REGION Network 2: Adress_Capa
         L     #Capa_Actual;
         L     1;
         -I;
         L     #Length_Capas;
         *I;
         L     #Offset_Capas;
         +I;
         T     #Adress_Capa;
END_REGION

REGION Network 3: Adress_Filas_DB
   New_Fil:NOP   0;
         L     #Índice_Filas;
         L     1;
         -I;
         L     #Length_Filas_DB;
         *I;
         L     #Offset_Filas_DB;
         +I;
         L     #Adress_Capa;
         +I;
         SLD   3;
         T     #Adress_Filas_DB_bit;
END_REGION

REGION Network 4: Adress_Filas_DI
         L     #Índice_Filas;
         L     1;
         -I;
         L     #Length_Filas_DI;
         *I;
         L     #Offset_Filas_DI;
         +I;
         T     #Adress_Filas_DI;
END_REGION

REGION Network 5: Adress_Elementos_DB
   New_Ele:NOP   0;
         L     #Índice_Elementos;
         L     1;
         -I;
         L     #Length_Elementos_DB_bit;
         *I;
         L     #Offset_Elementos_DB_bit;
         +I;
         L     #Adress_Filas_DB_bit;
         +I;
         T     #Adress_Elementos_DB_bit;
END_REGION

REGION Network 6: Adress_Elementos_DI
         L     #Índice_Elementos;
         L     1;
         -I;
         L     #Length_Elementos_DI;
         *I;
         L     #Offset_Elementos_DI;
         +I;
         L     #Adress_Filas_DI;
         +I;
         T     #Adress_Elementos_DI;
END_REGION

REGION Network 7: AR1 y AR2
         L     #Adress_Elementos_DB_bit;
         LAR1;
         L     #Adress_Elementos_DI;
         SLD   3;
         LAR2;
END_REGION

REGION Network 8: Transferencia de Figuras
   // No debería entrar nunca en este segmento, ya que necesita a Editando_Recetas y no entraría al bloque
         A     "Editando_Recetas";
         AN    "flanco"."nHMI.Pls_Inc_Capa";
         AN    "flanco"."nHMI.Pls_Dec_Capa";
         JCN   Fin;
         OPN   "DB_Receta_Actual";
         OPNDI "DB_Animación";
   // 0 = Invisible
   // 1 = V
   // 2 = H
   // 3 = HH
   //... Creo...
         L     DIB [ AR2 , P#0.0 ];
         L     0;
         ==I;
         JCN   NO_00;
         R     DBX[AR1,P#0.0];
         R     DBX [ AR1 , P#2.0 ];
         JU    Fin;
   NO_00:L     DIB [ AR2 , P#0.0 ];
         L     1;
         ==I;
         JCN   NO_10;
         S     DBX [ AR1 , P#0.0 ];
         R     DBX [ AR1 , P#2.0 ];
         JU    Fin;
   NO_10:L     DIB [ AR2 , P#0.0 ];
         L     2;
         ==I;
         JCN   NO_20;
         R     DBX[AR1,P#0.0];
         S     DBX [ AR1 , P#2.0 ];
         JU    Fin;
   NO_20:S     DBX [ AR1 , P#0.0 ];
         S     DBX [ AR1 , P#2.0 ];
   Fin:  NOP   0;
END_REGION

REGION Network 9: Transferencia de Figuras
   // En base a las figuras en bits de la receta actual, dibuja la capa gráficamente.
         OPN   "DB_Receta_Actual";
         OPNDI "DB_Animación";
   // 0 = Invisible
   // 1 = V
   // 2 = H
   // 3 = HH
   //... Creo...

         AN    DBX [ AR1 , P#0.0 ];
         AN    DBX [ AR1 , P#2.0 ];
         JCN   NO_0;
         L     0;
         JU    Transferir;
   NO_0: A     DBX [ AR1 , P#0.0 ];
         AN    DBX [ AR1 , P#2.0 ];
         JCN   NO_1;
         L     1;
         JU    Transferir;
   NO_1: AN    DBX [ AR1 , P#0.0 ];
         A     DBX [ AR1 , P#2.0 ];
         JCN   NO_2;
         L     2;
         JU    Transferir;
   NO_2: L     3;
   Transferir:T     DIB [ AR2 , P#0.0 ];
END_REGION

REGION Network 10: Transferencia de Elemento_SEL [ Anulado ]
   // Entra a veces en este segmento, se puede pulsar este botón dela pantalla 20 ó 21 [21 no entra al FC]
         A     "flanco"."pHMI.Pls_CargarReceta";
         JCN   Anular;
         OPN   "DB_Receta_Actual";
         OPNDI "DB_Animación";

         SET;
         A     DBX [ AR1 , P#4.0 ];
         JCN   otro;
         L     #Índice_Filas;
         T     "DB_Animación".Fila_SEL;
         L     #Índice_Elementos;
         T     "DB_Animación".Elemento_SEL;
   otro: NOP   0;

   Anular:NOP   0;
         OPN   "DB_Receta_Actual";
         OPNDI "DB_Animación";
END_REGION

REGION Network 11: Bucle Elementos
         L     #Índice_Elementos;
         L     1;
         +I;
         T     #Índice_Elementos;
         L     #Max_Nro_Elementos;
         <=I;
         JC    New_Ele;
END_REGION

REGION Network 12: Bucle Filas
         L     1;
         T     #Índice_Elementos;
         L     #Índice_Filas;
         L     1;
         +I;
         T     #Índice_Filas;
         L     #Max_Nro_Filas;
         <=I;
         JC    New_Fil;
END_REGION

REGION Network 13: Fin de Bloque
         BEU;
END_REGION
END_FUNCTION

FUNCTION "FC_INC_ELEM_ACTUAL" : Void   // FC19, STL
{ S7_Optimized_Access := 'FALSE' }
VERSION : 0.1
BEGIN

REGION Network 1: Constantes
         L     "Proceso Dosificador".Cant_Pallets;
         T     #Nro_Pallet;
         L     "Proceso Dosificador".Capa_Actual;
         T     #Capa_Actual;
         L     38;
         T     #Length_Capas;
         L     54;
         T     #Offset_Capas;
         L     6;
         T     #Length_Filas_DB;
         L     0;
         T     #Offset_Filas_DB;
         L     1;
         T     #Length_Elementos_DB_bit;
         L     0;
         T     #Offset_Elementos_DB_bit;

         L     1;
         T     #Índice_Filas;
         T     #Índice_Elementos;

         L     "Puntero".Max_Nro_Elementos;
         T     #Max_Nro_Elementos;
         L     "Puntero".Max_Nro_Filas;
         T     #Max_Nro_Filas;
         L     "Puntero".Max_Nro_Capas;
         T     #Max_Nro_Capas;
END_REGION

REGION Network 2: Adress_Capa
         L     #Capa_Actual;
         L     1;
         -I;
         L     #Length_Capas;
         *I;
         L     #Offset_Capas;
         +I;
         T     #Adress_Capa;
END_REGION

REGION Network 3: Adress_Filas
   New_Fil:NOP   0;
         L     #Índice_Filas;
         L     1;
         -I;
         L     #Length_Filas_DB;
         *I;
         L     #Offset_Filas_DB;
         +I;
         L     #Adress_Capa;
         +I;
         SLD   3;
         T     #Adress_Filas_DB_bit;
END_REGION

REGION Network 4: Adress_Elementos_DB
   New_Ele:NOP   0;
         L     #Índice_Elementos;
         L     1;
         -I;
         L     #Length_Elementos_DB_bit;
         *I;
         L     #Offset_Elementos_DB_bit;
         +I;
         L     #Adress_Filas_DB_bit;
         +I;
         T     #Adress_Elementos_DB_bit;
END_REGION

REGION Network 5: AR1
         L     #Adress_Elementos_DB_bit;
         LAR1;
END_REGION

REGION Network 6: Habilita ir 1 lugar a la IZQ si gráficamente existe un elemento a la izq.
         OPN   "DB_Receta_Actual";
         SET;
         R     #Habil_1_IZQ;
         L     #Índice_Elementos;
         L     #Max_Nro_Elementos;
         >=I;
         JC    No1IZQ;
         TAR1  AR2;
         L     1;
         +AR2;
         O     DBX [ AR2 , P#0.0 ];
         O     DBX [ AR2 , P#2.0 ];
         =     #Habil_1_IZQ;
   No1IZQ:NOP   0;
END_REGION

REGION Network 7: Habilita ir 2 lugar a la IZQ si gráficamente existen dos elementos a la izq.
         OPN   "DB_Receta_Actual";
         SET;
         R     #Habil_2_IZQ;
         L     #Índice_Elementos;
         L     1;
         +I;
         L     #Max_Nro_Elementos;
         >=I;
         JC    No2IZQ;
         TAR1  AR2;
         L     2;
         +AR2;
         O     DBX [ AR2 , P#0.0 ];
         O     DBX [ AR2 , P#2.0 ];
         =     #Habil_2_IZQ;
   No2IZQ:NOP   0;
END_REGION

REGION Network 8: Habilita ir a ABA_Elem_1 si gráficamente existe el primer elemento de la fila de abajo.
         OPN   "DB_Receta_Actual";
         SET;
         R     #Habil_1_ABA;
         L     #Índice_Filas;
         L     #Max_Nro_Filas;
         >=I;
         JC    No1ABA;
         L     #Adress_Filas_DB_bit;
         SRD   3;
         L     #Length_Filas_DB;
         +I;
         SLD   3;
         L     #Offset_Elementos_DB_bit;
         +I;
         LAR2;
         O     DBX [AR2, P#0.0];
         O     DBX [ AR2 , P#2.0 ];
         =     #Habil_1_ABA;
   No1ABA:NOP   0;
END_REGION

REGION Network 9: Habilita ir a ABA_Elem_2 si gráficamente existe el segundo elemento de la fila de abajo.
         OPN   "DB_Receta_Actual";
         SET;
         R     #Habil_2_ABA;
         L     #Índice_Filas;
         L     #Max_Nro_Filas;
         >=I;
         JC    No2ABA;
         L     #Adress_Filas_DB_bit;
         SRD   3;
         L     #Length_Filas_DB;
         +I;
         SLD   3;
         L     #Offset_Elementos_DB_bit;
         +I;
         L     #Length_Elementos_DB_bit;
         +I;
         LAR2;
         O     DBX [AR2, P#0.0];
         O     DBX [ AR2 , P#2.0 ];
         =     #Habil_2_ABA;
   No2ABA:NOP   0;
END_REGION

REGION Network 10: Habilita cambiar de CAPA_Elem_1, si existe el primer elemento de la próx. capa.
         OPN   "DB_Receta_Actual";
         SET;
         R     #Habil_1_CAPA;
         L     #Capa_Actual;
         L     #Max_Nro_Capas;
         >=I;
         JC    No1CAPA;
         L     #Adress_Capa;
         L     #Length_Capas;
         +I;
         L     #Offset_Filas_DB;
         +I;
         SLD   3;
         L     #Offset_Elementos_DB_bit;
         +I;
         LAR2;
         O     DBX [AR2, P#0.0];
         O     DBX [ AR2 , P#2.0 ];
         =     #Habil_1_CAPA;
   No1CAPA:NOP   0;
END_REGION

REGION Network 11: Habilita cambiar de CAPA_Elem_2, si existe el segundo elemento de la próx. capa.
         OPN   "DB_Receta_Actual";
         SET;
         R     #Habil_2_CAPA;
         L     #Capa_Actual;
         L     #Max_Nro_Capas;
         >=I;
         JC    No2CAPA;
         L     #Adress_Capa;
         L     #Length_Capas;
         +I;
         L     #Offset_Filas_DB;
         +I;
         SLD   3;
         L     #Offset_Elementos_DB_bit;
         +I;
         L     #Length_Elementos_DB_bit;
         +I;
         LAR2;
         O     DBX [AR2, P#0.0];
         O     DBX [ AR2 , P#2.0 ];
         =     #Habil_2_CAPA;
   No2CAPA:NOP   0;
END_REGION

REGION Network 12: #Elemento_Actual
         OPN   "DB_Receta_Actual";

         A     DBX [ AR1 , P#4.0 ];
         =     #Elemento_Actual;

         A     #Elemento_Actual;
         JCN   NoActual;
         TAR1  AR2;
END_REGION

REGION Network 13: NUM = 1
         L     #NUM;
         L     1;
         ==I;
         JCN   NUM_2;
         R     DBX [ AR1 , P#4.0 ];
         A     #Habil_1_IZQ;
         JCN   No_1_IZQ;

         TAR1  AR2;
         L     1;
         +AR2;
         S     DBX [ AR2 , P#4.0 ];
         JU    Fin;

   No_1_IZQ:A     #Habil_1_ABA;
         JCN   No_ABA;
         L     #Adress_Filas_DB_bit;
         SRD   3;
         L     #Length_Filas_DB;
         +I;
         SLD   3;
         L     #Offset_Elementos_DB_bit;
         +I;
         LAR2;
         SET;
         S     DBX [ AR2 , P#4.0 ];
         JU    Fin;

   No_ABA:A     #Habil_1_CAPA;
         JCN   No_CAPA;
         L     #Adress_Capa;
         L     #Length_Capas;
         +I;
         L     #Offset_Filas_DB;
         +I;
         SLD   3;
         L     #Offset_Elementos_DB_bit;
         +I;
         LAR2;
         S     DBX [ AR2 , P#4.0 ];
         L     #Capa_Actual;
         L     1;
         +I;
         T     #Capa_Actual;
         JU    Fin;

   No_CAPA:NOP   0;
         L     #Offset_Capas;
         L     #Offset_Filas_DB;
         +I;
         SLD   3;
         L     #Offset_Elementos_DB_bit;
         +I;
         LAR2;
         S     DBX [ AR2 , P#4.0 ];
         L     1;
         T     #Capa_Actual;
         L     #Nro_Pallet;
         L     1;
         +I;
         T     #Nro_Pallet;
         JU    Fin;
END_REGION

REGION Network 14: NUM = 2
   NUM_2:L     #NUM;
         L     2;
         ==I;
         JCN   NoNUM;
         R     DBX [ AR1 , P#4.0 ];
         A     #Habil_2_IZQ;
         JC    x_2IZQ;
         A     #Habil_1_IZQ;
         A     #Habil_1_ABA;
         JC    x_1IZQ_1ABA;
         A     #Habil_1_IZQ;
         A     #Habil_1_CAPA;
         JC    x_1IZQ_1CAPA;
         A     #Habil_1_IZQ;
         JC    x_1IZQ_1PALLET;
         A     #Habil_2_ABA;
         JC    x_2ABA;
         A     #Habil_1_ABA;
         A     #Habil_1_CAPA;
         JC    x_1ABA_1CAPA;
         A     #Habil_1_ABA;
         JC    x_1ABA_1PALLET;
         A     #Habil_2_CAPA;
         JC    x_2CAPA;
         A     #Habil_1_CAPA;
         JC    x_1CAPA_1PALLET;
         JU    x_2PALLET;

   x_2IZQ:NOP   0;
         TAR1  AR2;
         L     2;
         +AR2;
         S     DBX [ AR2 , P#4.0 ];
         JU    Fin;

   x_1IZQ_1ABA:NOP   0;
         L     #Adress_Filas_DB_bit;
         SRD   3;
         L     #Length_Filas_DB;
         +I;
         SLD   3;
         L     #Offset_Elementos_DB_bit;
         +I;
         LAR2;
         S     DBX [ AR2 , P#4.0 ];
         JU    Fin;

   x_2ABA:NOP   0;
         L     #Adress_Filas_DB_bit;
         SRD   3;
         L     #Length_Filas_DB;
         +I;
         SLD   3;
         L     #Offset_Elementos_DB_bit;
         +I;
         L     #Length_Elementos_DB_bit;
         +I;
         LAR2;
         S     DBX [ AR2 , P#4.0 ];
         JU    Fin;

   x_1IZQ_1CAPA:NOP   0;
   x_1ABA_1CAPA:NOP   0;
         L     #Adress_Capa;
         L     #Length_Capas;
         +I;
         L     #Offset_Filas_DB;
         +I;
         SLD   3;
         L     #Offset_Elementos_DB_bit;
         +I;
         LAR2;
         S     DBX [ AR2 , P#4.0 ];
         L     #Capa_Actual;
         L     1;
         +I;
         T     #Capa_Actual;
         JU    Fin;

   x_2CAPA:NOP   0;
         L     #Adress_Capa;
         L     #Length_Capas;
         +I;
         L     #Offset_Filas_DB;
         +I;
         SLD   3;
         L     #Offset_Elementos_DB_bit;
         +I;
         L     #Length_Elementos_DB_bit;
         +I;
         LAR2;
         S     DBX [ AR2 , P#4.0 ];
         L     #Capa_Actual;
         L     1;
         +I;
         T     #Capa_Actual;
         JU    Fin;

   x_1IZQ_1PALLET:NOP   0;
   x_1ABA_1PALLET:NOP   0;
   x_1CAPA_1PALLET:NOP   0;
         L     #Offset_Capas;
         L     #Offset_Filas_DB;
         +I;
         SLD   3;
         L     #Offset_Elementos_DB_bit;
         +I;
         LAR2;
         S     DBX [ AR2 , P#4.0 ];
         L     1;
         T     #Capa_Actual;
         L     #Nro_Pallet;
         L     1;
         +I;
         T     #Nro_Pallet;
         JU    Fin;

   x_2PALLET:NOP   0;
         L     #Offset_Capas;
         L     #Offset_Filas_DB;
         +I;
         SLD   3;
         L     #Offset_Elementos_DB_bit;
         +I;
         L     #Length_Elementos_DB_bit;
         +I;
         LAR2;
         S     DBX [ AR2 , P#4.0 ];
         L     1;
         T     #Capa_Actual;
         L     #Nro_Pallet;
         L     1;
         +I;
         T     #Nro_Pallet;
         JU    Fin;
END_REGION

REGION Network 15: No elemento actual
   NoNUM:JU    Fin;
   NoActual:NOP   0;
END_REGION

REGION Network 16: Bucle Elementos
         L     #Índice_Elementos;
         L     1;
         +I;
         T     #Índice_Elementos;
         L     #Max_Nro_Elementos;
         <=I;
         JC    New_Ele;
END_REGION

REGION Network 17: Bucle Filas
         L     1;
         T     #Índice_Elementos;
         L     #Índice_Filas;
         L     1;
         +I;
         T     #Índice_Filas;
         L     #Max_Nro_Filas;
         <=I;
         JC    New_Fil;
END_REGION

REGION Network 18: #Error
         SET;
         S     #Error;
         JU    ERROR;
END_REGION

REGION Network 19: Fin de Bloque
   Fin:  SET;
         R     #Error;
         OPN   "DB_Receta_Actual";
         AN    DBX [ AR2 , P#0.0 ];
         AN    DBX [ AR2 , P#2.0 ];
         JCN   NO_0;
         L     0;
         JU    Transferir;
   NO_0: A     DBX [ AR2 , P#0.0 ];
         AN    DBX [ AR2 , P#2.0 ];
         JCN   NO_1;
         L     1;
         JU    Transferir;
   NO_1: AN    DBX [ AR2 , P#0.0 ];
         A     DBX [ AR2 , P#2.0 ];
         JCN   NO_2;
         L     2;
         JU    Transferir;
   NO_2: L     3;
   Transferir:T     "Proceso Dosificador".Elemento_Actual;
   // 0 = Invisible
   // 1 = V
   // 2 = H
   // 3 = HH


   ERROR:L     #Capa_Actual;
         T     "Proceso Dosificador".Capa_Actual;
         L     #Nro_Pallet;
         T     "Proceso Dosificador".Cant_Pallets;
END_REGION
END_FUNCTION

FUNCTION "FC_Ver_Recetas_faltaEditar" : Void   // FC21, STL
TITLE = Muestra los datos de la receta seleccionada
{ S7_Optimized_Access := 'FALSE' }
VERSION : 0.1
BEGIN

REGION Network 1: Constantes
         L     "Puntero".Offset_Recetas;
         T     #Offset_Recetas;
         L     "Puntero".Length_Recetas;
         T     #Length_Recetas;
         L     "Puntero".Offset_Nombre_Receta;
         T     #Offset_Nombre_Receta_DB;
         L     "Puntero".Max_Nro_Recetas;
         T     #Max_Nro_Recetas;
   //
         L     "Puntero".Offset_CapasDist_Receta;
   //    L     51
         T     #Offset_CapasDist_Receta_DB;
         L     "Puntero".Offset_CantCapas_Receta;
   //    L     50
         T     #Offset_CantCapas_Receta_DB;
         L     "Puntero".Length_Nombre_Receta;
   //    L     50
         T     #Length_Nombre_Receta;
   //
         L     316;
         T     #Offset_CantCapas_Receta_DI;
         L     317;
         T     #Offset_CapasDist_Receta_DI;
   //
         L     "DB_Animación".Nro_Receta_Edición;
         T     #Nro_Receta;
   //
         A     "flanco"."nHMI.Pls_Inc_Receta";
         =     #fn_Inc_Receta;
         A     "flanco"."nHMI.Pls_Dec_Receta";
         =     #fn_Dec_Receta;
   //
         L     "HMI".Imagen_Actual;
         T     #Imagen;
END_REGION

REGION Network 2
         L     #Nro_Receta;
         L     #Max_Nro_Recetas;
         <I;
         A     #fn_Inc_Receta;
         JCN   noINC;
         TAK;
         L     1;
         +I;
         JU    Transferir;
   noINC:NOP   0;

         L     #Nro_Receta;
         L     1;
         >I;
         A     #fn_Dec_Receta;
         JCN   noDEC;
         TAK;
         L     1;
         -I;
         JU    Transferir;
   noDEC:NOP   0;
         L     #Nro_Receta;
   Transferir:T     #Nro_Receta;
END_REGION

REGION Network 3: Abrir la receta correspondiente
         L     #Nro_Receta;
         L     1;
         -I;
         L     #Length_Recetas;
         *I;
         L     #Offset_Recetas;
         +I;
         T     #Adress_Receta;
END_REGION

REGION Network 4: Transferir Nombre de receta
         OPN   "DB_RECETAS";
         OPNDI "DB_Animación";
         L     #Adress_Receta;
         L     #Offset_Nombre_Receta_DB;
         +I;
         SLD   3;
         LAR1;
         L     266;
         SLD   3;
         LAR2;
         L     0;
         T     #K;
   Bucle:SLD   3;
         +AR1;
         +AR2;

         A     "Editando_Recetas";
         JCN   NoEsc_0;
         L     DIB [ AR2 , P#0.0 ];
         T     DBB [ AR1 , P#0.0 ];
   NoEsc_0:NOP   0;

         L     DBB [ AR1 , P#0.0 ];
         T     DIB [ AR2 , P#0.0 ];
         L     #K;
         L     1;
         +I;
         T     #K;
         L     #Length_Nombre_Receta;
         <I;
         L     1;
         JC    Bucle;
END_REGION

REGION Network 5: Transferir Número de capas por pallet
         OPN   "DB_RECETAS";
         OPNDI "DB_Animación";
         L     #Adress_Receta;
         L     #Offset_CantCapas_Receta_DB;
         +I;
         SLD   3;
         LAR1;
         L     #Offset_CantCapas_Receta_DI;
         SLD   3;
         LAR2;

         A     "Editando_Recetas";
         JCN   NoEsc_1;
         L     DIB [ AR2 , P#0.0 ];
         T     DBB [ AR1 , P#0.0 ];
   NoEsc_1:NOP   0;

         L     DBB [AR1, P#0.0];
         T     DIB [ AR2 , P#0.0 ];
END_REGION

REGION Network 6: Transferir Número de capas distintas
         OPN   "DB_RECETAS";
         OPNDI "DB_Animación";
         L     #Adress_Receta;
         L     #Offset_CapasDist_Receta_DB;
         +I;
         SLD   3;
         LAR1;
         L     #Offset_CapasDist_Receta_DI;
         SLD   3;
         LAR2;

         A     "Editando_Recetas";
         JCN   NoEsc_2;
         L     DIB [ AR2 , P#0.0 ];
         T     DBB [ AR1 , P#0.0 ];
   NoEsc_2:NOP   0;

         L     DBB [AR1, P#0.0];
         T     DIB [ AR2 , P#0.0 ];
END_REGION

REGION Network 7
         L     #Nro_Receta;
         T     "DB_Animación".Nro_Receta_Edición;
END_REGION
END_FUNCTION

FUNCTION "FC_RESET_ELEM_ACTUAL" : Void   // FC22, STL
{ S7_Optimized_Access := 'FALSE' }
VERSION : 0.1
// Con los datos del dosificador, setea el bit de elemento actual en DB_Receta_Actual
BEGIN

REGION Network 1: Constantes
         L     "Proceso Empujador".Capa_Actual;
         T     #Capa_Empuj;
         L     "Proceso Dosificador".Cant_Pallets;
         T     #Nro_Pallet;
         L     "Proceso Dosificador".Capa_Actual;
         T     #Capa_Actual;
         L     38;
         T     #Length_Capas;
         L     54;
         T     #Offset_Capas;
         L     6;
         T     #Length_Filas_DB;
         L     0;
         T     #Offset_Filas_DB;
         L     1;
         T     #Length_Elementos_DB_bit;
         L     0;
         T     #Offset_Elementos_DB_bit;

         L     1;
         T     #Índice_Capas;
         T     #Índice_Filas;
         T     #Índice_Elementos;

         L     "Puntero".Max_Nro_Elementos;
         T     #Max_Nro_Elementos;
         L     "Puntero".Max_Nro_Filas;
         T     #Max_Nro_Filas;
         L     "Puntero".Max_Nro_Capas;
         T     #Max_Nro_Capas;

         L     "DB_Animación".Fila_SEL;
         T     #Fila_SEL;
         L     "DB_Animación".Elemento_SEL;
         T     #Elemento_SEL;
END_REGION

REGION Network 2: Set CAPA
         OPN   "DB_Receta_Actual";
   //     SPA   no
         L     #Capa_Empuj;
         T     #Capa_Actual;
   no:   NOP   0;
END_REGION

REGION Network 3: Adress_Capa
   New_Cap:L     #Índice_Capas;
         L     1;
         -I;
         L     #Length_Capas;
         *I;
         L     #Offset_Capas;
         +I;
         T     #Adress_Capa;
END_REGION

REGION Network 4: Adress_Filas
   New_Fil:L     #Índice_Filas;
         L     1;
         -I;
         L     #Length_Filas_DB;
         *I;
         L     #Offset_Filas_DB;
         +I;
         L     #Adress_Capa;
         +I;
         SLD   3;
         T     #Adress_Filas_DB_bit;
END_REGION

REGION Network 5: Adress_Elementos_DB
   New_Ele:L     #Índice_Elementos;
         L     1;
         -I;
         L     #Length_Elementos_DB_bit;
         *I;
         L     #Offset_Elementos_DB_bit;
         +I;
         L     #Adress_Filas_DB_bit;
         +I;
         T     #Adress_Elementos_DB_bit;
END_REGION

REGION Network 6: AR1
         L     #Adress_Elementos_DB_bit;
         LAR1;
END_REGION

REGION Network 7: SR Elemento actual
   //  SPA   end
         L     #Capa_Actual;
         L     #Índice_Capas;
         ==I;
         JCN   noSEL;
         L     #Fila_SEL;
         L     #Índice_Filas;
         ==I;
         JCN   noSEL;
         L     #Elemento_SEL;
         L     #Índice_Elementos;
         ==I;
         JCN   noSEL;
         SET;
         S     DBX [AR1,P#4.0];
         JU    end;
   noSEL:SET;
         R     DBX [ AR1 , P#4.0 ];
   end:  NOP   0;
END_REGION

REGION Network 8: Bucle Elementos
         L     #Índice_Elementos;
         L     1;
         +I;
         T     #Índice_Elementos;
         L     #Max_Nro_Elementos;
         <=I;
         JC    New_Ele;
END_REGION

REGION Network 9: Bucle Filas
         L     1;
         T     #Índice_Elementos;
         L     #Índice_Filas;
         L     1;
         +I;
         T     #Índice_Filas;
         L     #Max_Nro_Filas;
         <=I;
         JC    New_Fil;
END_REGION

REGION Network 10: Bucle Capas
         L     1;
         T     #Índice_Filas;
         L     #Índice_Capas;
         L     1;
         +I;
         T     #Índice_Capas;
         L     #Max_Nro_Capas;
         <=I;
         JC    New_Cap;
END_REGION

REGION Network 11: Fin de Bloque
         L     #Capa_Actual;
         T     "Proceso Dosificador".Capa_Actual;
         L     #Nro_Pallet;
         T     "Proceso Dosificador".Cant_Pallets;
END_REGION
END_FUNCTION

(* ===== HMI "HMI_RT_1" =====
connection "Conexión_HMI_1": ETHERNET, SIMATIC S7 300/400 MPI

HMI tags "Tabla de variables estándar"
   "Elemento_1" : Int, internal
   "Elemento_2" : Int, internal
   "Elemento_3" : Int, internal
   "DB_Animación_Nro_Receta_Edición" : Byte, 1 s
   "DB_Animación_Nombre_Receta_Edición" : Array [0..49] of Char, 1 s
   "DB_Animación_Capas_X_Pallet_Edición" : Byte, 1 s
   "DB_Animación_CapasDistintas_Edición" : Byte, 1 s
   "VerCartel_TerminarPallet" : Bool, internal
   "PLC a HMI_Almacén_Pallets" : Bool, 1 s
   "PLC a HMI_Elevador" : Bool, 1 s
   "PLC a HMI_Seg_Elevador" : Bool, 1 s
   "PLC a HMI_Transp_2" : Bool, 1 s
   "PLC a HMI_Transp_3" : Bool, 1 s
   "PLC a HMI_Transp_4" : Bool, 1 s
   "PLC a HMI_Transp_5" : Bool, 1 s
   "PLC a HMI_Descarga" : Bool, 1 s
   "PLC a HMI_Avance_1_2" : Bool, 1 s
   "PLC a HMI_Avance_2_3" : Bool, 1 s
   "PLC a HMI_Avance_3_4" : Bool, 1 s
   "PLC a HMI_Avance_5_Desc" : Bool, 1 s
   "PLC a HMI_Avance_4_5" : Bool, 1 s
   "PLC a HMI_PEDIDO_ENVOLV" : Bool, 1 s
   "PLC a HMI_ENVOLVER" : Bool, 1 s
   "PLC a HMI_PALLET_ENVUELTO" : Bool, 1 s
   "PLC a HMI_ETIQUETAR" : Bool, 1 s
   "PLC a HMI_CICLO_OK" : Bool, 1 s
   "PLC a HMI_HOME_PISTON" : Bool, 100 ms
   "ALARMAS_1" : Word, 1 s
   "ALARMAS_2" : Word, 1 s
   "ALARMAS_3" : Word, 1 s
   "ALARMAS_4" : Word, 1 s
   "ALARMAS_5" : Word, 1 s
   "ALARMAS_6" : Word, 1 s
   "ALARMAS_7" : Word, 1 s
   "Pallet_Transporte1_a_Transporte2" : Bool = PLC "Pallet_Transporte1_a_Transporte2", 1 s
   "Pallet_Transporte2_a_Envolvedora" : Bool = PLC "Pallet_Transporte2_a_Envolvedora", 1 s
   "Pallet_Envolvedora_a_Etiquetadora" : Bool = PLC "Pallet_Envolvedora_a_Etiquetadora", 1 s
   "Pallet_Etiquetadora_a_Transporte5" : Bool = PLC "Pallet_Etiquetadora_a_Transporte5", 1 s
   "Pallet_Transporte5_a_Descarga" : Bool = PLC "Pallet_Transporte5_a_Descarga", 1 s
   "Sin_Ala" : Bool = PLC "Sin_Ala", 1 s
   "HMI_TP1_a_TP2" : Bool, 1 s
   "HMI_TP2_a_TP3" : Bool, 1 s
   "HMI_TP3_a_TP4" : Bool, 1 s
   "HMI_TP4_a_TP5" : Bool, 1 s
   "HMI_TP5_a_Desc" : Bool, 1 s
   "Brazo_Descarga_Man" : Bool = PLC "Brazo_Descarga_Man", 1 s
   "iSnsBarrDesc_Atr" : Bool = PLC "iSnsBarrDesc_Atr", 1 s
   "iSnsAscen_Arr" : Bool = PLC "iSnsAscen_Arr", 1 s
   "iSnsAscen_Aba_Len" : Bool = PLC "iSnsAscen_Aba_Len", 1 s
   "iSnsAscen_Aba_Par" : Bool = PLC "iSnsAscen_Aba_Par", 1 s
   "iSnsPlataf_Ade" : Bool = PLC "iSnsPlataf_Ade", 1 s
   "iSnsPlataf_Atr" : Bool = PLC "iSnsPlataf_Atr", 1 s
   "iSnsRetEmpuBrazo" : Bool = PLC "iSnsRetEmpuBrazo", 1 s
   "iSnsEmpj_Arriba" : Bool = PLC "iSnsEmpj_Arriba", 1 s
   "iSnsEmpj_Abajo" : Bool = PLC "iSnsEmpj_Abajo", 1 s
   "iSnsEmpj_Ade_Par" : Bool = PLC "iSnsEmpj_Ade_Par", 1 s
   "iSnsEmpj_Ade_Len" : Bool = PLC "iSnsEmpj_Ade_Len", 1 s
   "iSnsEmpj_Atr_Len" : Bool = PLC "iSnsEmpj_Atr_Len", 1 s
   "iSnsEmpj_Atr_Par" : Bool = PLC "iSnsEmpj_Atr_Par", 1 s
   "iSnsEmpj_MedCamin" : Bool = PLC "iSnsEmpj_MedCamin", 1 s
   "iSnsCajaEn_21.22" : Bool = PLC "iSnsCajaEn_21.22", 1 s
   "iSnsCajaEn_21.26" : Bool = PLC "iSnsCajaEn_21.26", 1 s
   "oTransp_21.10" : Bool = PLC "oTransp_21.10", 1 s
   "oTransp_21.22" : Bool = PLC "oTransp_21.22", 1 s
   "oTransp_21.24" : Bool = PLC "oTransp_21.24", 1 s
   "oTransp_21.26" : Bool = PLC "oTransp_21.26", 1 s
   "Color_Alarmas" : Byte = PLC "Color_Alarmas", 1 s
   "DB_Animación_Capa_Actual_Edición" : Byte, 1 s
   "DB_Velocidades_Dosif_LímInf_Vel" : Real, 1 s
   "DB_Velocidades_Dosif_Vel_Ráp" : Real, 1 s
   "DB_Velocidades_Dosif_LímSup_Vel" : Real, 1 s
   "DB_Velocidades_Ascens_LímInf_Vel" : Real, 1 s
   "DB_Velocidades_Ascens_VelRáp_Arr" : Real, 1 s
   "DB_Velocidades_Ascens_VelLen_Arr" : Real, 1 s
   "DB_Velocidades_Ascens_VelRáp_Aba" : Real, 1 s
   "DB_Velocidades_Ascens_VelLen_Aba" : Real, 1 s
   "DB_Velocidades_Ascens_LímSup_Vel" : Real, 1 s
   "DB_Velocidades_Empuj_LímInf_Vel" : Real, 1 s
   "DB_Velocidades_Empuj_VelRáp_Ade" : Real, 1 s
   "DB_Velocidades_Empuj_VelLen_Ade" : Real, 1 s
   "DB_Velocidades_Empuj_VelRáp_Atr" : Real, 1 s
   "DB_Velocidades_Empuj_VelLen_Atr" : Real, 1 s
   "DB_Velocidades_Empuj_LímSup_Vel" : Real, 1 s
   "HMI_Pls_Inc_Figura_Sel" : Bool, 1 s
   "HMI_Pls_Inc_Capa_Editando" : Bool, 1 s
   "HMI_Pls_Dec_Capa_Editando" : Bool, 1 s
   "DB_Animación_Usar_Pistón" : Bool, 1 s
   "Siempre_1" : Bool, internal
   "ALARMAS_8" : Word, 1 s
   "HMI_Cartones_1_o_2" : Bool, 1 s
   "Siempre_0" : Bool, internal
   "DB_Carton_Manual_Catoneo_Manual_Hab" : Bool, 1 s
   "DB_Carton_Manual_CM_FrenoCiclo" : Bool, 1 s
   "HMI_hab_etiq" : Bool, 1 s
   "HMI_hab_fechadora1" : Bool, 1 s
   "HMI_hab_fechadora2" : Bool, 1 s

HMI tags "PLC_a_HMI"
   "PLC_a_HMI_Fila[1].Offset_Y" : Int, 100 ms
   "PLC_a_HMI_Fila[1].Elemento[1].Figura" : Byte, 100 ms
   "PLC_a_HMI_Fila[1].Elemento[1].Offset_X" : Int, 100 ms
   "PLC_a_HMI_Fila[1].Elemento[1].Estado" : Byte, 100 ms
   "PLC_a_HMI_Fila[1].Elemento[2].Figura" : Byte, 100 ms
   "PLC_a_HMI_Fila[1].Elemento[2].Offset_X" : Int, 100 ms
   "PLC_a_HMI_Fila[1].Elemento[2].Estado" : Byte, 100 ms
   "PLC_a_HMI_Fila[1].Elemento[3].Figura" : Byte, 100 ms
   "PLC_a_HMI_Fila[1].Elemento[3].Offset_X" : Int, 100 ms
   "PLC_a_HMI_Fila[1].Elemento[3].Estado" : Byte, 100 ms
   "PLC_a_HMI_Fila[1].Elemento[4].Figura" : Byte, 100 ms
   "PLC_a_HMI_Fila[1].Elemento[4].Offset_X" : Int, 100 ms
   "PLC_a_HMI_Fila[1].Elemento[4].Estado" : Byte, 100 ms
   "PLC_a_HMI_Fila[1].Elemento[5].Figura" : Byte, 100 ms
   "PLC_a_HMI_Fila[1].Elemento[5].Offset_X" : Int, 100 ms
   "PLC_a_HMI_Fila[1].Elemento[5].Estado" : Byte, 100 ms
   "PLC_a_HMI_Fila[1].Elemento[6].Figura" : Byte, 100 ms
   "PLC_a_HMI_Fila[1].Elemento[6].Offset_X" : Int, 100 ms
   "PLC_a_HMI_Fila[1].Elemento[6].Estado" : Byte, 100 ms
   "PLC_a_HMI_Fila[1].Elemento[7].Figura" : Byte, 100 ms
   "PLC_a_HMI_Fila[1].Elemento[7].Offset_X" : Int, 100 ms
   "PLC_a_HMI_Fila[1].Elemento[7].Estado" : Byte, 100 ms
   "PLC_a_HMI_Fila[1].Elemento[8].Figura" : Byte, 100 ms
   "PLC_a_HMI_Fila[1].Elemento[8].Offset_X" : Int, 100 ms
   "PLC_a_HMI_Fila[1].Elemento[8].Estado" : Byte, 100 ms
   "PLC_a_HMI_Fila[1].Elemento[9].Figura" : Byte, 100 ms
   "PLC_a_HMI_Fila[1].Elemento[9].Offset_X" : Int, 100 ms
   "PLC_a_HMI_Fila[1].Elemento[9].Estado" : Byte, 100 ms
   "PLC_a_HMI_Fila[1].Elemento[10].Figura" : Byte, 100 ms
   "PLC_a_HMI_Fila[1].Elemento[10].Offset_X" : Int, 100 ms
   "PLC_a_HMI_Fila[1].Elemento[10].Estado" : Byte, 100 ms
   "PLC_a_HMI_Fila[2].Offset_Y" : Int, 100 ms
   "PLC_a_HMI_Fila[2].Elemento[1].Figura" : Byte, 100 ms
   "PLC_a_HMI_Fila[2].Elemento[1].Offset_X" : Int, 100 ms
   "PLC_a_HMI_Fila[2].Elemento[1].Estado" : Byte, 100 ms
   "PLC_a_HMI_Fila[2].Elemento[2].Figura" : Byte, 100 ms
   "PLC_a_HMI_Fila[2].Elemento[2].Offset_X" : Int, 100 ms
   "PLC_a_HMI_Fila[2].Elemento[2].Estado" : Byte, 100 ms
   "PLC_a_HMI_Fila[2].Elemento[3].Figura" : Byte, 100 ms
   "PLC_a_HMI_Fila[2].Elemento[3].Offset_X" : Int, 100 ms
   "PLC_a_HMI_Fila[2].Elemento[3].Estado" : Byte, 100 ms
   "PLC_a_HMI_Fila[2].Elemento[4].Figura" : Byte, 100 ms
   "PLC_a_HMI_Fila[2].Elemento[4].Offset_X" : Int, 100 ms
   "PLC_a_HMI_Fila[2].Elemento[4].Estado" : Byte, 100 ms
   "PLC_a_HMI_Fila[2].Elemento[5].Figura" : Byte, 100 ms
   "PLC_a_HMI_Fila[2].Elemento[5].Offset_X" : Int, 100 ms
   "PLC_a_HMI_Fila[2].Elemento[5].Estado" : Byte, 100 ms
   "PLC_a_HMI_Fila[2].Elemento[6].Figura" : Byte, 100 ms
   "PLC_a_HMI_Fila[2].Elemento[6].Offset_X" : Int, 100 ms
   "PLC_a_HMI_Fila[2].Elemento[6].Estado" : Byte, 100 ms
   "PLC_a_HMI_Fila[2].Elemento[7].Figura" : Byte, 100 ms
   "PLC_a_HMI_Fila[2].Elemento[7].Offset_X" : Int, 100 ms
   "PLC_a_HMI_Fila[2].Elemento[7].Estado" : Byte, 100 ms
   "PLC_a_HMI_Fila[2].Elemento[8].Figura" : Byte, 100 ms
   "PLC_a_HMI_Fila[2].Elemento[8].Offset_X" : Int, 100 ms
   "PLC_a_HMI_Fila[2].Elemento[8].Estado" : Byte, 100 ms
   "PLC_a_HMI_Fila[2].Elemento[9].Figura" : Byte, 100 ms
   "PLC_a_HMI_Fila[2].Elemento[9].Offset_X" : Int, 100 ms
   "PLC_a_HMI_Fila[2].Elemento[9].Estado" : Byte, 100 ms
   "PLC_a_HMI_Fila[2].Elemento[10].Figura" : Byte, 100 ms
   "PLC_a_HMI_Fila[2].Elemento[10].Offset_X" : Int, 100 ms
   "PLC_a_HMI_Fila[2].Elemento[10].Estado" : Byte, 100 ms
   "PLC_a_HMI_Fila[3].Offset_Y" : Int, 100 ms
   "PLC_a_HMI_Fila[3].Elemento[1].Figura" : Byte, 100 ms
   "PLC_a_HMI_Fila[3].Elemento[1].Offset_X" : Int, 100 ms
   "PLC_a_HMI_Fila[3].Elemento[1].Estado" : Byte, 100 ms
   "PLC_a_HMI_Fila[3].Elemento[2].Figura" : Byte, 100 ms
   "PLC_a_HMI_Fila[3].Elemento[2].Offset_X" : Int, 100 ms
   "PLC_a_HMI_Fila[3].Elemento[2].Estado" : Byte, 100 ms
   "PLC_a_HMI_Fila[3].Elemento[3].Figura" : Byte, 100 ms
   "PLC_a_HMI_Fila[3].Elemento[3].Offset_X" : Int, 100 ms
   "PLC_a_HMI_Fila[3].Elemento[3].Estado" : Byte, 100 ms
   "PLC_a_HMI_Fila[3].Elemento[4].Figura" : Byte, 100 ms
   "PLC_a_HMI_Fila[3].Elemento[4].Offset_X" : Int, 100 ms
   "PLC_a_HMI_Fila[3].Elemento[4].Estado" : Byte, 100 ms
   "PLC_a_HMI_Fila[3].Elemento[5].Figura" : Byte, 100 ms
   "PLC_a_HMI_Fila[3].Elemento[5].Offset_X" : Int, 100 ms
   "PLC_a_HMI_Fila[3].Elemento[5].Estado" : Byte, 100 ms
   "PLC_a_HMI_Fila[3].Elemento[6].Figura" : Byte, 100 ms
   "PLC_a_HMI_Fila[3].Elemento[6].Offset_X" : Int, 100 ms
   "PLC_a_HMI_Fila[3].Elemento[6].Estado" : Byte, 100 ms
   "PLC_a_HMI_Fila[3].Elemento[7].Figura" : Byte, 100 ms
   "PLC_a_HMI_Fila[3].Elemento[7].Offset_X" : Int, 100 ms
   "PLC_a_HMI_Fila[3].Elemento[7].Estado" : Byte, 100 ms
   "PLC_a_HMI_Fila[3].Elemento[8].Figura" : Byte, 100 ms
   "PLC_a_HMI_Fila[3].Elemento[8].Offset_X" : Int, 100 ms
   "PLC_a_HMI_Fila[3].Elemento[8].Estado" : Byte, 100 ms
   "PLC_a_HMI_Fila[3].Elemento[9].Figura" : Byte, 100 ms
   "PLC_a_HMI_Fila[3].Elemento[9].Offset_X" : Int, 100 ms
   "PLC_a_HMI_Fila[3].Elemento[9].Estado" : Byte, 100 ms
   "PLC_a_HMI_Fila[3].Elemento[10].Figura" : Byte, 100 ms
   "PLC_a_HMI_Fila[3].Elemento[10].Offset_X" : Int, 100 ms
   "PLC_a_HMI_Fila[3].Elemento[10].Estado" : Byte, 100 ms
   "PLC_a_HMI_Fila[4].Offset_Y" : Int, 100 ms
   "PLC_a_HMI_Fila[4].Elemento[1].Figura" : Byte, 100 ms
   "PLC_a_HMI_Fila[4].Elemento[1].Offset_X" : Int, 100 ms
   "PLC_a_HMI_Fila[4].Elemento[1].Estado" : Byte, 100 ms
   "PLC_a_HMI_Fila[4].Elemento[2].Figura" : Byte, 100 ms
   "PLC_a_HMI_Fila[4].Elemento[2].Offset_X" : Int, 100 ms
   "PLC_a_HMI_Fila[4].Elemento[2].Estado" : Byte, 100 ms
   "PLC_a_HMI_Fila[4].Elemento[3].Figura" : Byte, 100 ms
   "PLC_a_HMI_Fila[4].Elemento[3].Offset_X" : Int, 100 ms
   "PLC_a_HMI_Fila[4].Elemento[3].Estado" : Byte, 100 ms
   "PLC_a_HMI_Fila[4].Elemento[4].Figura" : Byte, 100 ms
   "PLC_a_HMI_Fila[4].Elemento[4].Offset_X" : Int, 100 ms
   "PLC_a_HMI_Fila[4].Elemento[4].Estado" : Byte, 100 ms
   "PLC_a_HMI_Fila[4].Elemento[5].Figura" : Byte, 100 ms
   "PLC_a_HMI_Fila[4].Elemento[5].Offset_X" : Int, 100 ms
   "PLC_a_HMI_Fila[4].Elemento[5].Estado" : Byte, 100 ms
   "PLC_a_HMI_Fila[4].Elemento[6].Figura" : Byte, 100 ms
   "PLC_a_HMI_Fila[4].Elemento[6].Offset_X" : Int, 100 ms
   "PLC_a_HMI_Fila[4].Elemento[6].Estado" : Byte, 100 ms
   "PLC_a_HMI_Fila[4].Elemento[7].Figura" : Byte, 100 ms
   "PLC_a_HMI_Fila[4].Elemento[7].Offset_X" : Int, 100 ms
   "PLC_a_HMI_Fila[4].Elemento[7].Estado" : Byte, 100 ms
   "PLC_a_HMI_Fila[4].Elemento[8].Figura" : Byte, 100 ms
   "PLC_a_HMI_Fila[4].Elemento[8].Offset_X" : Int, 100 ms
   "PLC_a_HMI_Fila[4].Elemento[8].Estado" : Byte, 100 ms
   "PLC_a_HMI_Fila[4].Elemento[9].Figura" : Byte, 100 ms
   "PLC_a_HMI_Fila[4].Elemento[9].Offset_X" : Int, 100 ms
   "PLC_a_HMI_Fila[4].Elemento[9].Estado" : Byte, 100 ms
   "PLC_a_HMI_Fila[4].Elemento[10].Figura" : Byte, 100 ms
   "PLC_a_HMI_Fila[4].Elemento[10].Offset_X" : Int, 100 ms
   "PLC_a_HMI_Fila[4].Elemento[10].Estado" : Byte, 100 ms
   "PLC_a_HMI_Fila[5].Offset_Y" : Int, 100 ms
   "PLC_a_HMI_Fila[5].Elemento[1].Figura" : Byte, 100 ms
   "PLC_a_HMI_Fila[5].Elemento[1].Offset_X" : Int, 100 ms
   "PLC_a_HMI_Fila[5].Elemento[1].Estado" : Byte, 100 ms
   "PLC_a_HMI_Fila[5].Elemento[2].Figura" : Byte, 100 ms
   "PLC_a_HMI_Fila[5].Elemento[2].Offset_X" : Int, 100 ms
   "PLC_a_HMI_Fila[5].Elemento[2].Estado" : Byte, 100 ms
   "PLC_a_HMI_Fila[5].Elemento[3].Figura" : Byte, 100 ms
   "PLC_a_HMI_Fila[5].Elemento[3].Offset_X" : Int, 100 ms
   "PLC_a_HMI_Fila[5].Elemento[3].Estado" : Byte, 100 ms
   "PLC_a_HMI_Fila[5].Elemento[4].Figura" : Byte, 100 ms
   "PLC_a_HMI_Fila[5].Elemento[4].Offset_X" : Int, 100 ms
   "PLC_a_HMI_Fila[5].Elemento[4].Estado" : Byte, 100 ms
   "PLC_a_HMI_Fila[5].Elemento[5].Figura" : Byte, 100 ms
   "PLC_a_HMI_Fila[5].Elemento[5].Offset_X" : Int, 100 ms
   "PLC_a_HMI_Fila[5].Elemento[5].Estado" : Byte, 100 ms
   "PLC_a_HMI_Fila[5].Elemento[6].Figura" : Byte, 100 ms
   "PLC_a_HMI_Fila[5].Elemento[6].Offset_X" : Int, 100 ms
   "PLC_a_HMI_Fila[5].Elemento[6].Estado" : Byte, 100 ms
   "PLC_a_HMI_Fila[5].Elemento[7].Figura" : Byte, 100 ms
   "PLC_a_HMI_Fila[5].Elemento[7].Offset_X" : Int, 100 ms
   "PLC_a_HMI_Fila[5].Elemento[7].Estado" : Byte, 100 ms
   "PLC_a_HMI_Fila[5].Elemento[8].Figura" : Byte, 100 ms
   "PLC_a_HMI_Fila[5].Elemento[8].Offset_X" : Int, 100 ms
   "PLC_a_HMI_Fila[5].Elemento[8].Estado" : Byte, 100 ms
   "PLC_a_HMI_Fila[5].Elemento[9].Figura" : Byte, 100 ms
   "PLC_a_HMI_Fila[5].Elemento[9].Offset_X" : Int, 100 ms
   "PLC_a_HMI_Fila[5].Elemento[9].Estado" : Byte, 100 ms
   "PLC_a_HMI_Fila[5].Elemento[10].Figura" : Byte, 100 ms
   "PLC_a_HMI_Fila[5].Elemento[10].Offset_X" : Int, 100 ms
   "PLC_a_HMI_Fila[5].Elemento[10].Estado" : Byte, 100 ms
   "PLC_a_HMI_Fila[6].Offset_Y" : Int, 100 ms
   "PLC_a_HMI_Fila[6].Elemento[1].Figura" : Byte, 100 ms
   "PLC_a_HMI_Fila[6].Elemento[1].Offset_X" : Int, 100 ms
   "PLC_a_HMI_Fila[6].Elemento[1].Estado" : Byte, 100 ms
   "PLC_a_HMI_Fila[6].Elemento[2].Figura" : Byte, 100 ms